// TIA Portal project "Respirator2020_V16" (V16) (continued)
REGION Network 5: Peep Supervisor
   RUNG wire#powerrail
      "VariableSupervisor_DB_Peep"(SetpointIncrement := "OperatingParameters".PeepPBPlus, SetpointDecrement := "OperatingParameters".PeepPBMinus, Max := 50.0, Min := 3.0, SetpointMax := "OperatingParameters".PeepMax, SetpointMin := "OperatingParameters".PeepMin, InOutSetpoint := "OperatingParameters".PeepSetpoint, InOutAlarmHI := "ProcessData".PeepSetpointAlarmHI, InOutPreAlarmHI := "ProcessData".PeepSetpointPreAlarmHI, InOutAlarmLOW := "ProcessData".PeepSetpointAlarmLOW, InOutPreAlarmLOW := "ProcessData".PeepSetpointPreAlarmLOW)
   END_RUNG
   // the same network as SCL:
   "VariableSupervisor_DB_Peep"(SetpointIncrement := "OperatingParameters".PeepPBPlus,   // "VariableSupervisor"
                           SetpointDecrement := "OperatingParameters".PeepPBMinus,
                           Max := 50.0,
                           Min := 3.0,
                           SetpointMax := "OperatingParameters".PeepMax,
                           SetpointMin := "OperatingParameters".PeepMin,
                           InOutSetpoint := "OperatingParameters".PeepSetpoint,
                           InOutAlarmHI := "ProcessData".PeepSetpointAlarmHI,
                           InOutPreAlarmHI := "ProcessData".PeepSetpointPreAlarmHI,
                           InOutAlarmLOW := "ProcessData".PeepSetpointAlarmLOW,
                           InOutPreAlarmLOW := "ProcessData".PeepSetpointPreAlarmLOW);
END_REGION

REGION Network 6: Frequency Supervisor
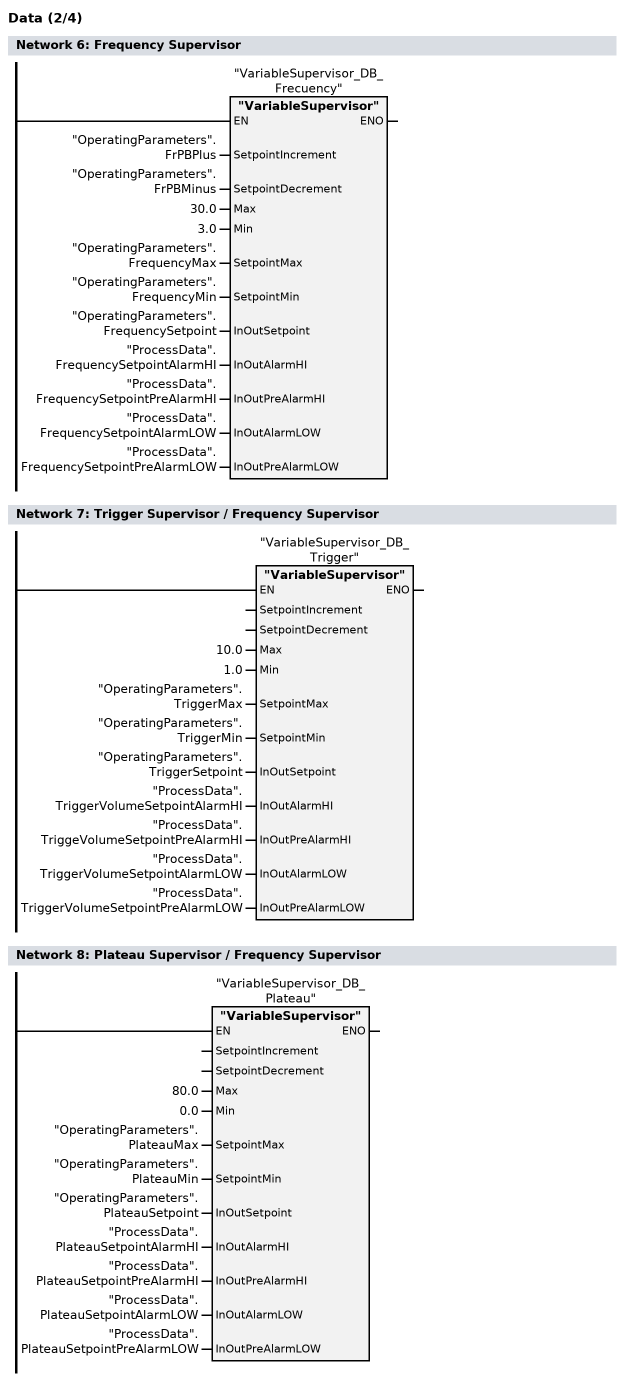
   RUNG wire#powerrail
      "VariableSupervisor_DB_Frecuency"(SetpointIncrement := "OperatingParameters".FrPBPlus, SetpointDecrement := "OperatingParameters".FrPBMinus, Max := 30.0, Min := 3.0, SetpointMax := "OperatingParameters".FrequencyMax, SetpointMin := "OperatingParameters".FrequencyMin, InOutSetpoint := "OperatingParameters".FrequencySetpoint, InOutAlarmHI := "ProcessData".FrequencySetpointAlarmHI, InOutPreAlarmHI := "ProcessData".FrequencySetpointPreAlarmHI, InOutAlarmLOW := "ProcessData".FrequencySetpointAlarmLOW, InOutPreAlarmLOW := "ProcessData".FrequencySetpointPreAlarmLOW)
   END_RUNG
   // the same network as SCL:
   "VariableSupervisor_DB_Frecuency"(SetpointIncrement := "OperatingParameters".FrPBPlus,   // "VariableSupervisor"
                           SetpointDecrement := "OperatingParameters".FrPBMinus,
                           Max := 30.0,
                           Min := 3.0,
                           SetpointMax := "OperatingParameters".FrequencyMax,
                           SetpointMin := "OperatingParameters".FrequencyMin,
                           InOutSetpoint := "OperatingParameters".FrequencySetpoint,
                           InOutAlarmHI := "ProcessData".FrequencySetpointAlarmHI,
                           InOutPreAlarmHI := "ProcessData".FrequencySetpointPreAlarmHI,
                           InOutAlarmLOW := "ProcessData".FrequencySetpointAlarmLOW,
                           InOutPreAlarmLOW := "ProcessData".FrequencySetpointPreAlarmLOW);
END_REGION

REGION Network 7: Trigger Supervisor / Frequency Supervisor
   RUNG wire#powerrail
      "VariableSupervisor_DB_Trigger"(SetpointIncrement :=, SetpointDecrement :=, Max := 10.0, Min := 1.0, SetpointMax := "OperatingParameters".TriggerMax, SetpointMin := "OperatingParameters".TriggerMin, InOutSetpoint := "OperatingParameters".TriggerSetpoint, InOutAlarmHI := "ProcessData".TriggerVolumeSetpointAlarmHI, InOutPreAlarmHI := "ProcessData".TriggeVolumeSetpointPreAlarmHI, InOutAlarmLOW := "ProcessData".TriggerVolumeSetpointAlarmLOW, InOutPreAlarmLOW := "ProcessData".TriggerVolumeSetpointPreAlarmLOW)
   END_RUNG
   // the same network as SCL:
   "VariableSupervisor_DB_Trigger"(Max := 10.0,   // "VariableSupervisor"
                           Min := 1.0,
                           SetpointMax := "OperatingParameters".TriggerMax,
                           SetpointMin := "OperatingParameters".TriggerMin,
                           InOutSetpoint := "OperatingParameters".TriggerSetpoint,
                           InOutAlarmHI := "ProcessData".TriggerVolumeSetpointAlarmHI,
                           InOutPreAlarmHI := "ProcessData".TriggeVolumeSetpointPreAlarmHI,
                           InOutAlarmLOW := "ProcessData".TriggerVolumeSetpointAlarmLOW,
                           InOutPreAlarmLOW := "ProcessData".TriggerVolumeSetpointPreAlarmLOW);
END_REGION

REGION Network 8: Plateau Supervisor / Frequency Supervisor
   RUNG wire#powerrail
      "VariableSupervisor_DB_Plateau"(SetpointIncrement :=, SetpointDecrement :=, Max := 80.0, Min := 0.0, SetpointMax := "OperatingParameters".PlateauMax, SetpointMin := "OperatingParameters".PlateauMin, InOutSetpoint := "OperatingParameters".PlateauSetpoint, InOutAlarmHI := "ProcessData".PlateauSetpointAlarmHI, InOutPreAlarmHI := "ProcessData".PlateauSetpointPreAlarmHI, InOutAlarmLOW := "ProcessData".PlateauSetpointAlarmLOW, InOutPreAlarmLOW := "ProcessData".PlateauSetpointPreAlarmLOW)
   END_RUNG
   // the same network as SCL:
   "VariableSupervisor_DB_Plateau"(Max := 80.0,   // "VariableSupervisor"
                           Min := 0.0,
                           SetpointMax := "OperatingParameters".PlateauMax,
                           SetpointMin := "OperatingParameters".PlateauMin,
                           InOutSetpoint := "OperatingParameters".PlateauSetpoint,
                           InOutAlarmHI := "ProcessData".PlateauSetpointAlarmHI,
                           InOutPreAlarmHI := "ProcessData".PlateauSetpointPreAlarmHI,
                           InOutAlarmLOW := "ProcessData".PlateauSetpointAlarmLOW,
                           InOutPreAlarmLOW := "ProcessData".PlateauSetpointPreAlarmLOW);
END_REGION

REGION Network 9: TidalVolume Supervisor / Frequency Supervisor
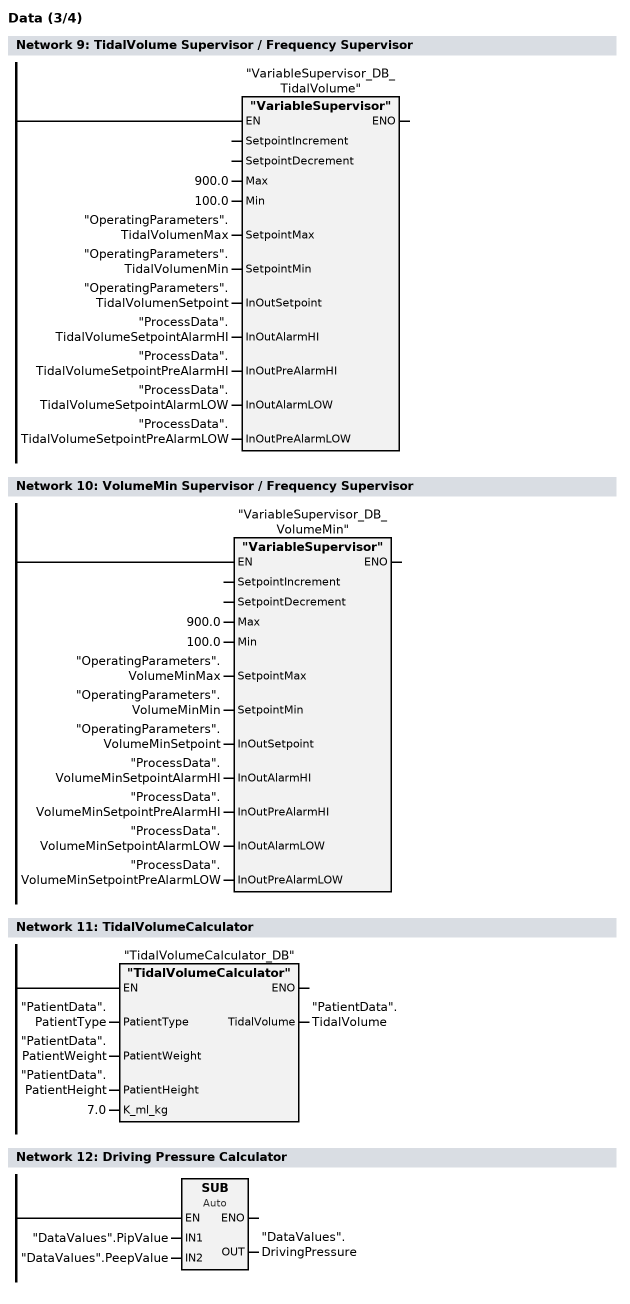
   RUNG wire#powerrail
      "VariableSupervisor_DB_TidalVolume"(SetpointIncrement :=, SetpointDecrement :=, Max := 900.0, Min := 100.0, SetpointMax := "OperatingParameters".TidalVolumenMax, SetpointMin := "OperatingParameters".TidalVolumenMin, InOutSetpoint := "OperatingParameters".TidalVolumenSetpoint, InOutAlarmHI := "ProcessData".TidalVolumeSetpointAlarmHI, InOutPreAlarmHI := "ProcessData".TidalVolumeSetpointPreAlarmHI, InOutAlarmLOW := "ProcessData".TidalVolumeSetpointAlarmLOW, InOutPreAlarmLOW := "ProcessData".TidalVolumeSetpointPreAlarmLOW)
   END_RUNG
   // the same network as SCL:
   "VariableSupervisor_DB_TidalVolume"(Max := 900.0,   // "VariableSupervisor"
                           Min := 100.0,
                           SetpointMax := "OperatingParameters".TidalVolumenMax,
                           SetpointMin := "OperatingParameters".TidalVolumenMin,
                           InOutSetpoint := "OperatingParameters".TidalVolumenSetpoint,
                           InOutAlarmHI := "ProcessData".TidalVolumeSetpointAlarmHI,
                           InOutPreAlarmHI := "ProcessData".TidalVolumeSetpointPreAlarmHI,
                           InOutAlarmLOW := "ProcessData".TidalVolumeSetpointAlarmLOW,
                           InOutPreAlarmLOW := "ProcessData".TidalVolumeSetpointPreAlarmLOW);
END_REGION

REGION Network 10: VolumeMin Supervisor / Frequency Supervisor
   RUNG wire#powerrail
      "VariableSupervisor_DB_VolumeMin"(SetpointIncrement :=, SetpointDecrement :=, Max := 900.0, Min := 100.0, SetpointMax := "OperatingParameters".VolumeMinMax, SetpointMin := "OperatingParameters".VolumeMinMin, InOutSetpoint := "OperatingParameters".VolumeMinSetpoint, InOutAlarmHI := "ProcessData".VolumeMinSetpointAlarmHI, InOutPreAlarmHI := "ProcessData".VolumeMinSetpointPreAlarmHI, InOutAlarmLOW := "ProcessData".VolumeMinSetpointAlarmLOW, InOutPreAlarmLOW := "ProcessData".VolumeMinSetpointPreAlarmLOW)
   END_RUNG
   // the same network as SCL:
   "VariableSupervisor_DB_VolumeMin"(Max := 900.0,   // "VariableSupervisor"
                           Min := 100.0,
                           SetpointMax := "OperatingParameters".VolumeMinMax,
                           SetpointMin := "OperatingParameters".VolumeMinMin,
                           InOutSetpoint := "OperatingParameters".VolumeMinSetpoint,
                           InOutAlarmHI := "ProcessData".VolumeMinSetpointAlarmHI,
                           InOutPreAlarmHI := "ProcessData".VolumeMinSetpointPreAlarmHI,
                           InOutAlarmLOW := "ProcessData".VolumeMinSetpointAlarmLOW,
                           InOutPreAlarmLOW := "ProcessData".VolumeMinSetpointPreAlarmLOW);
END_REGION

REGION Network 11: TidalVolumeCalculator
   RUNG wire#powerrail
      "TidalVolumeCalculator_DB"(PatientType := "PatientData".PatientType, PatientWeight := "PatientData".PatientWeight, PatientHeight := "PatientData".PatientHeight, K_ml_kg := 7.0, TidalVolume => "PatientData".TidalVolume)
   END_RUNG
   // the same network as SCL:
   "TidalVolumeCalculator_DB"(PatientType := "PatientData".PatientType,   // "TidalVolumeCalculator"
                           PatientWeight := "PatientData".PatientWeight,
                           PatientHeight := "PatientData".PatientHeight,
                           K_ml_kg := 7.0,
                           TidalVolume => "PatientData".TidalVolume);
END_REGION

REGION Network 12: Driving Pressure Calculator
   RUNG wire#powerrail
      Sub(in1 := "DataValues".PipValue, in2 := "DataValues".PeepValue, out => "DataValues".DrivingPressure)
   END_RUNG
   // the same network as SCL:
   "DataValues".DrivingPressure := "DataValues".PipValue - "DataValues".PeepValue;
END_REGION

REGION Network 13: Ratio Calculator
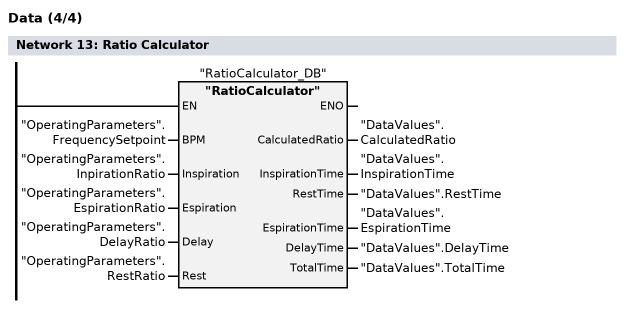
   RUNG wire#powerrail
      "RatioCalculator_DB"(BPM := "OperatingParameters".FrequencySetpoint, Inspiration := "OperatingParameters".InpirationRatio, Espiration := "OperatingParameters".EspirationRatio, Delay := "OperatingParameters".DelayRatio, Rest := "OperatingParameters".RestRatio, CalculatedRatio => "DataValues".CalculatedRatio, InspirationTime => "DataValues".InspirationTime, RestTime => "DataValues".RestTime, EspirationTime => "DataValues".EspirationTime, DelayTime => "DataValues".DelayTime, TotalTime => "DataValues".TotalTime)
   END_RUNG
   // the same network as SCL:
   "RatioCalculator_DB"(BPM := "OperatingParameters".FrequencySetpoint,   // "RatioCalculator"
                        Inspiration := "OperatingParameters".InpirationRatio,
                        Espiration := "OperatingParameters".EspirationRatio,
                        Delay := "OperatingParameters".DelayRatio,
                        Rest := "OperatingParameters".RestRatio,
                        CalculatedRatio => "DataValues".CalculatedRatio,
                        InspirationTime => "DataValues".InspirationTime,
                        RestTime => "DataValues".RestTime,
                        EspirationTime => "DataValues".EspirationTime,
                        DelayTime => "DataValues".DelayTime,
                        TotalTime => "DataValues".TotalTime);
END_REGION
END_FUNCTION_BLOCK

FUNCTION_BLOCK "TidalVolumeCalculator"   // FB11, SCL
{ S7_Optimized_Access := 'TRUE' }
AUTHOR : JL_Cristobal_2020
VERSION : 0.1
   VAR_INPUT
      PatientType : Int;
      PatientWeight : Real;
      PatientHeight : Real;
      K_ml_kg : Real;
   END_VAR
   VAR_OUTPUT
      TidalVolume : Real;
   END_VAR
   VAR
      CorrectedWeight : Real;
   END_VAR
BEGIN
   //**************************************************************************************************
   // TidalVolumeCalculator
   //**************************************************************************************************

   // Sex Selection
   CASE #PatientType OF
       1:  // Man
           #CorrectedWeight := 50.0;
       2:  // Woman
           #CorrectedWeight := 45.5;
       ELSE  // Not selected
           #CorrectedWeight := 0.0;;
   END_CASE;

   // Calc
   IF #CorrectedWeight <> 0 THEN
       #TidalVolume:= #K_ml_kg *((#CorrectedWeight+0.91)*(#PatientHeight));
       ELSE
           #TidalVolume := 0.0;
   END_IF;
END_FUNCTION_BLOCK

// folder: 2_SensorComm

FUNCTION_BLOCK "SensorComm_PtP_Freeport"   // FB20, SCL
{ S7_Optimized_Access := 'FALSE' }
AUTHOR : JL_Cristobal_2020
VERSION : 0.1
   VAR_OUTPUT
      OutputStatus : Struct
         Pressure1 : Real;
         Pressure2 : Real;
         VolumeAccumulated : Real;
         Flow : Real;
         TEMPERATURA_SONICA_PROMEDIO : Real;
         TEMPERATURA_PT100 : Real;
         HUMEDAD_RELATIVA : Real;
         PRESION_ATMOSFERICA : Real;
         DIRECCION_BRUJULA : Real;
         RADIACION_SOLAR : Real;
         VEL_PROMEDIO_VIENTO : Real;
         DIR_MEDIA_VIENTO : Real;
         HUMEDAD_ABSOLUTA : Real;
         PUNTO_ROCIO : Real;
         DIRECCION_VIENTO_GRADOS : Real;
         VEL_VIENTO_EJE_V : Real;
         VEL_VIENTO_EJE_U : Real;
         ERROR_MEDICION_VELOCIDAD : Bool;
         ERROR_MEDICION_BRUJULA : Bool;
         ERROR_MEDICION_TEMPERATURA : Bool;
         ERROR_MEDICION_HUMEDAD : Bool;
         ERROR_MEDICION_PRESION : Bool;
         ERROR_MEDICION_RADIACION_SOLAR : Bool;
      END_STRUCT;
      Pressure1 : Real;
      Pressure2 : Real;
      VolumeAccumulated : Real;
      Flow : Real;
      ErrorPressure1 : Bool;
      ErrorPressure2 : Bool;
      ErrorVolumeAccumulated : Bool;
      ErrorFlow : Bool;
   END_VAR
   VAR
      InputData : Struct
         Config_REQ : Bool;
         Reset_REQ : Bool;
      END_STRUCT;
      OutputData : Struct
         Config_DONE : Bool;
         Config_ERROR : Bool;
         Config_STAT : Word;
         Reset_DONE : Bool;
         Reset_ERROR : Bool;
         Reset_STAT : Word;
         Receive_P2P_NDR : Bool;
         Receive_P2P_ERROR : Bool;
         Receive_P2P_STAT : Word;
         Receive_P2P_Length : Word;
         Send_P2P_DONE : Bool;
         Send_P2P_ERROR : Bool;
         Send_P2P_STAT : Word;
      END_STRUCT;
      Control : Struct
         While_Section : Bool;
         COM_RST : Bool;
         Config_ERROR_save : Word;
         Reset_ERROR_save : Word;
         P2P_ERROR_save : Word;
         P2P_NDR_save : Word;
         Rcv_Length_save : Int;
      END_STRUCT;
      RecvBuffer : Array[1..254] of Byte;
      TransBuffer : Array[1..254] of Byte;
      IntermediateData : Struct
         Pressure1 : String;
         Pressure2 : String;
         VolumeAccumulated : String;
         Flow : String;
         Errors : String;
      END_STRUCT;
   END_VAR
BEGIN
   //**************************************************************************************************
   // Reading STATUS
   //**************************************************************************************************
   IF TRUE THEN
       // Pressure-1
       Chars_TO_Strg(Chars := "SensorComm_C_buffer_ptp".Ringbuffer,
                     pChars := 2,
                     Cnt := 6,
                     Strg => #IntermediateData.Pressure1);
       STRG_VAL(IN := #IntermediateData.Pressure1,
                FORMAT := W#16#0000,
                P := 1,
                OUT => #OutputStatus.Pressure1);
       #Pressure1 := #OutputStatus.Pressure1;

       // Pressure-2
       Chars_TO_Strg(Chars := "SensorComm_C_buffer_ptp".Ringbuffer,
                     pChars := 10,
                     Cnt := 6,
                     Strg => #IntermediateData.Pressure2);
       STRG_VAL(IN := #IntermediateData.Pressure2,
                FORMAT := W#16#0000,
                P := 1,
                OUT => #OutputStatus.Pressure2);
       #Pressure2 := #OutputStatus.Pressure2;

       // Volume Accumulated
       Chars_TO_Strg(Chars := "SensorComm_C_buffer_ptp".Ringbuffer,
                     pChars := 18,
                     Cnt := 6,
                     Strg => #IntermediateData.VolumeAccumulated);
       STRG_VAL(IN := #IntermediateData.VolumeAccumulated,
                FORMAT := W#16#0000,
                P := 1,
                OUT => #OutputStatus.VolumeAccumulated);
       #VolumeAccumulated := #OutputStatus.VolumeAccumulated;

       // Flow
       Chars_TO_Strg(Chars := "SensorComm_C_buffer_ptp".Ringbuffer,
                     pChars := 26,
                     Cnt := 6,
                     Strg => #IntermediateData.Flow);
       STRG_VAL(IN := #IntermediateData.Flow,
                FORMAT := W#16#0000,
                P := 1,
                OUT => #OutputStatus.Flow);
       #Flow := #OutputStatus.Flow;

        // Errors
       Chars_TO_Strg(Chars := "SensorComm_C_buffer_ptp".Ringbuffer,
                     pChars := 74,
                     Cnt := 6,
                     Strg => #IntermediateData.Errors);
   END_IF;
END_FUNCTION_BLOCK

// folder: 3_Alarms

FUNCTION_BLOCK "Alarms"   // FB5, LAD
TITLE = Alarms, Packing and Transport to HMI
{ S7_Optimized_Access := 'TRUE' }
AUTHOR : JL_Cristobal_2020
VERSION : 0.1
   VAR_IN_OUT
      AlarmsPack0 : Bool;
      AlarmsPack1 : Bool;
      AlarmsPack2 : Bool;
      AlarmsPack3 : Bool;
   END_VAR
BEGIN

REGION Network 1: Peak Alarms
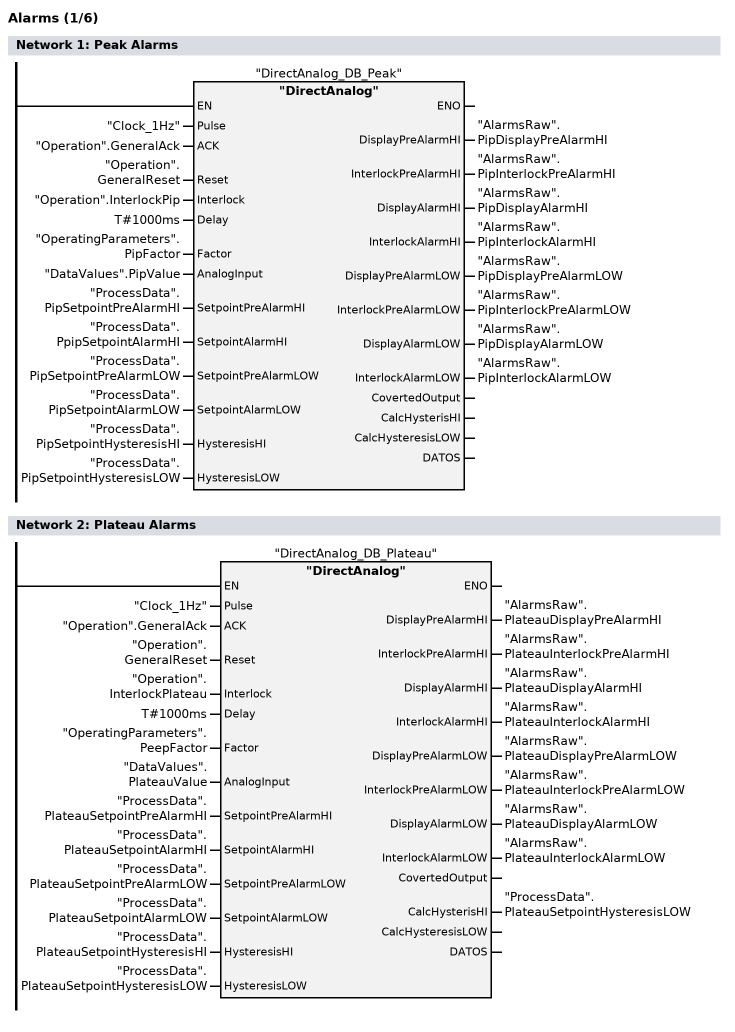
   RUNG wire#powerrail
      "DirectAnalog_DB_Peak"(Pulse := "Clock_1Hz", ACK := "Operation".GeneralAck, Reset := "Operation".GeneralReset, Interlock := "Operation".InterlockPip, Delay := T#1000ms, Factor := "OperatingParameters".PipFactor, AnalogInput := "DataValues".PipValue, SetpointPreAlarmHI := "ProcessData".PipSetpointPreAlarmHI, SetpointAlarmHI := "ProcessData".PpipSetpointAlarmHI, SetpointPreAlarmLOW := "ProcessData".PipSetpointPreAlarmLOW, SetpointAlarmLOW := "ProcessData".PipSetpointAlarmLOW, HysteresisHI := "ProcessData".PipSetpointHysteresisHI, HysteresisLOW := "ProcessData".PipSetpointHysteresisLOW, DisplayPreAlarmHI => "AlarmsRaw".PipDisplayPreAlarmHI, InterlockPreAlarmHI => "AlarmsRaw".PipInterlockPreAlarmHI, DisplayAlarmHI => "AlarmsRaw".PipDisplayAlarmHI, InterlockAlarmHI => "AlarmsRaw".PipInterlockAlarmHI, DisplayPreAlarmLOW => "AlarmsRaw".PipDisplayPreAlarmLOW, InterlockPreAlarmLOW => "AlarmsRaw".PipInterlockPreAlarmLOW, DisplayAlarmLOW => "AlarmsRaw".PipDisplayAlarmLOW, InterlockAlarmLOW => "AlarmsRaw".PipInterlockAlarmLOW, CovertedOutput =>, CalcHysterisHI =>, CalcHysteresisLOW =>, DATOS =>)
   END_RUNG
   // the same network as SCL:
   "DirectAnalog_DB_Peak"(Pulse := "Clock_1Hz",   // "DirectAnalog"
                          ACK := "Operation".GeneralAck,
                          Reset := "Operation".GeneralReset,
                          Interlock := "Operation".InterlockPip,
                          Delay := T#1000ms,
                          Factor := "OperatingParameters".PipFactor,
                          AnalogInput := "DataValues".PipValue,
                          SetpointPreAlarmHI := "ProcessData".PipSetpointPreAlarmHI,
                          SetpointAlarmHI := "ProcessData".PpipSetpointAlarmHI,
                          SetpointPreAlarmLOW := "ProcessData".PipSetpointPreAlarmLOW,
                          SetpointAlarmLOW := "ProcessData".PipSetpointAlarmLOW,
                          HysteresisHI := "ProcessData".PipSetpointHysteresisHI,
                          HysteresisLOW := "ProcessData".PipSetpointHysteresisLOW,
                          DisplayPreAlarmHI => "AlarmsRaw".PipDisplayPreAlarmHI,
                          InterlockPreAlarmHI => "AlarmsRaw".PipInterlockPreAlarmHI,
                          DisplayAlarmHI => "AlarmsRaw".PipDisplayAlarmHI,
                          InterlockAlarmHI => "AlarmsRaw".PipInterlockAlarmHI,
                          DisplayPreAlarmLOW => "AlarmsRaw".PipDisplayPreAlarmLOW,
                          InterlockPreAlarmLOW => "AlarmsRaw".PipInterlockPreAlarmLOW,
                          DisplayAlarmLOW => "AlarmsRaw".PipDisplayAlarmLOW,
                          InterlockAlarmLOW => "AlarmsRaw".PipInterlockAlarmLOW);
END_REGION

REGION Network 2: Plateau Alarms
   RUNG wire#powerrail
      "DirectAnalog_DB_Plateau"(Pulse := "Clock_1Hz", ACK := "Operation".GeneralAck, Reset := "Operation".GeneralReset, Interlock := "Operation".InterlockPlateau, Delay := T#1000ms, Factor := "OperatingParameters".PeepFactor, AnalogInput := "DataValues".PlateauValue, SetpointPreAlarmHI := "ProcessData".PlateauSetpointPreAlarmHI, SetpointAlarmHI := "ProcessData".PlateauSetpointAlarmHI, SetpointPreAlarmLOW := "ProcessData".PlateauSetpointPreAlarmLOW, SetpointAlarmLOW := "ProcessData".PlateauSetpointAlarmLOW, HysteresisHI := "ProcessData".PlateauSetpointHysteresisHI, HysteresisLOW := "ProcessData".PlateauSetpointHysteresisLOW, DisplayPreAlarmHI => "AlarmsRaw".PlateauDisplayPreAlarmHI, InterlockPreAlarmHI => "AlarmsRaw".PlateauInterlockPreAlarmHI, DisplayAlarmHI => "AlarmsRaw".PlateauDisplayAlarmHI, InterlockAlarmHI => "AlarmsRaw".PlateauInterlockAlarmHI, DisplayPreAlarmLOW => "AlarmsRaw".PlateauDisplayPreAlarmLOW, InterlockPreAlarmLOW => "AlarmsRaw".PlateauInterlockPreAlarmLOW, DisplayAlarmLOW => "AlarmsRaw".PlateauDisplayAlarmLOW, InterlockAlarmLOW => "AlarmsRaw".PlateauInterlockAlarmLOW, CovertedOutput =>, CalcHysterisHI => "ProcessData".PlateauSetpointHysteresisLOW, CalcHysteresisLOW =>, DATOS =>)
   END_RUNG
   // the same network as SCL:
   "DirectAnalog_DB_Plateau"(Pulse := "Clock_1Hz",   // "DirectAnalog"
                           ACK := "Operation".GeneralAck,
                           Reset := "Operation".GeneralReset,
                           Interlock := "Operation".InterlockPlateau,
                           Delay := T#1000ms,
                           Factor := "OperatingParameters".PeepFactor,
                           AnalogInput := "DataValues".PlateauValue,
                           SetpointPreAlarmHI := "ProcessData".PlateauSetpointPreAlarmHI,
                           SetpointAlarmHI := "ProcessData".PlateauSetpointAlarmHI,
                           SetpointPreAlarmLOW := "ProcessData".PlateauSetpointPreAlarmLOW,
                           SetpointAlarmLOW := "ProcessData".PlateauSetpointAlarmLOW,
                           HysteresisHI := "ProcessData".PlateauSetpointHysteresisHI,
                           HysteresisLOW := "ProcessData".PlateauSetpointHysteresisLOW,
                           DisplayPreAlarmHI => "AlarmsRaw".PlateauDisplayPreAlarmHI,
                           InterlockPreAlarmHI => "AlarmsRaw".PlateauInterlockPreAlarmHI,
                           DisplayAlarmHI => "AlarmsRaw".PlateauDisplayAlarmHI,
                           InterlockAlarmHI => "AlarmsRaw".PlateauInterlockAlarmHI,
                           DisplayPreAlarmLOW => "AlarmsRaw".PlateauDisplayPreAlarmLOW,
                           InterlockPreAlarmLOW => "AlarmsRaw".PlateauInterlockPreAlarmLOW,
                           DisplayAlarmLOW => "AlarmsRaw".PlateauDisplayAlarmLOW,
                           InterlockAlarmLOW => "AlarmsRaw".PlateauInterlockAlarmLOW,
                           CalcHysterisHI => "ProcessData".PlateauSetpointHysteresisLOW);
END_REGION

REGION Network 3: Peep Alarms
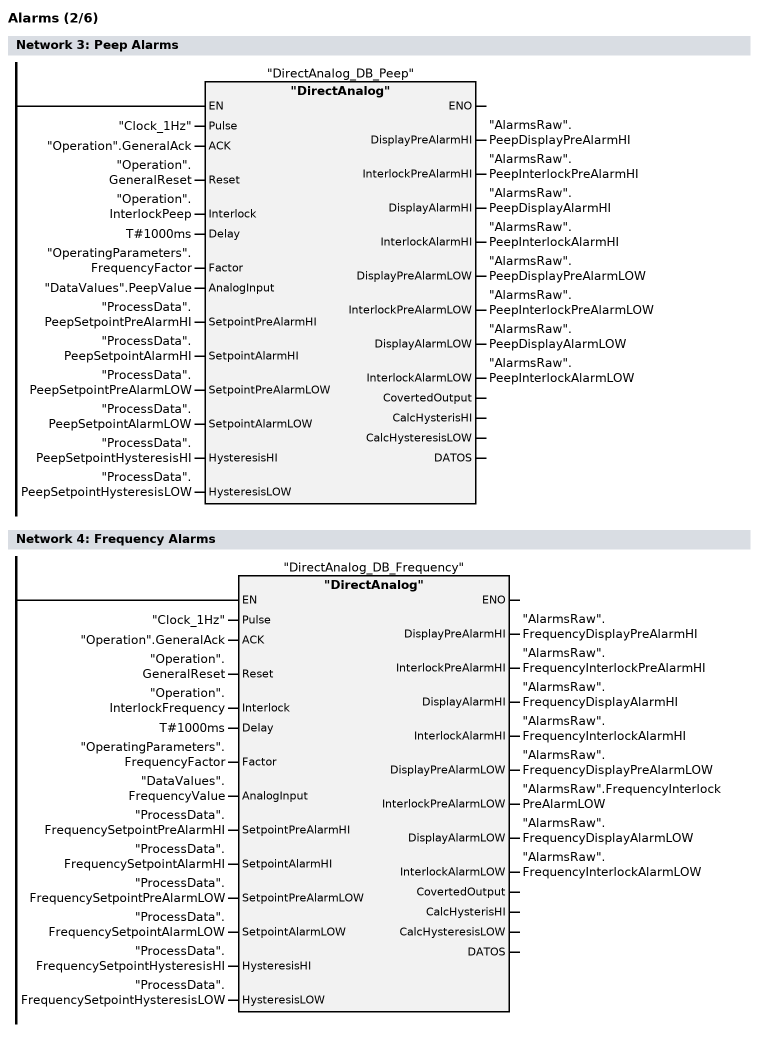
   RUNG wire#powerrail
      "DirectAnalog_DB_Peep"(Pulse := "Clock_1Hz", ACK := "Operation".GeneralAck, Reset := "Operation".GeneralReset, Interlock := "Operation".InterlockPeep, Delay := T#1000ms, Factor := "OperatingParameters".FrequencyFactor, AnalogInput := "DataValues".PeepValue, SetpointPreAlarmHI := "ProcessData".PeepSetpointPreAlarmHI, SetpointAlarmHI := "ProcessData".PeepSetpointAlarmHI, SetpointPreAlarmLOW := "ProcessData".PeepSetpointPreAlarmLOW, SetpointAlarmLOW := "ProcessData".PeepSetpointAlarmLOW, HysteresisHI := "ProcessData".PeepSetpointHysteresisHI, HysteresisLOW := "ProcessData".PeepSetpointHysteresisLOW, DisplayPreAlarmHI => "AlarmsRaw".PeepDisplayPreAlarmHI, InterlockPreAlarmHI => "AlarmsRaw".PeepInterlockPreAlarmHI, DisplayAlarmHI => "AlarmsRaw".PeepDisplayAlarmHI, InterlockAlarmHI => "AlarmsRaw".PeepInterlockAlarmHI, DisplayPreAlarmLOW => "AlarmsRaw".PeepDisplayPreAlarmLOW, InterlockPreAlarmLOW => "AlarmsRaw".PeepInterlockPreAlarmLOW, DisplayAlarmLOW => "AlarmsRaw".PeepDisplayAlarmLOW, InterlockAlarmLOW => "AlarmsRaw".PeepInterlockAlarmLOW, CovertedOutput =>, CalcHysterisHI =>, CalcHysteresisLOW =>, DATOS =>)
   END_RUNG
   // the same network as SCL:
   "DirectAnalog_DB_Peep"(Pulse := "Clock_1Hz",   // "DirectAnalog"
                          ACK := "Operation".GeneralAck,
                          Reset := "Operation".GeneralReset,
                          Interlock := "Operation".InterlockPeep,
                          Delay := T#1000ms,
                          Factor := "OperatingParameters".FrequencyFactor,
                          AnalogInput := "DataValues".PeepValue,
                          SetpointPreAlarmHI := "ProcessData".PeepSetpointPreAlarmHI,
                          SetpointAlarmHI := "ProcessData".PeepSetpointAlarmHI,
                          SetpointPreAlarmLOW := "ProcessData".PeepSetpointPreAlarmLOW,
                          SetpointAlarmLOW := "ProcessData".PeepSetpointAlarmLOW,
                          HysteresisHI := "ProcessData".PeepSetpointHysteresisHI,
                          HysteresisLOW := "ProcessData".PeepSetpointHysteresisLOW,
                          DisplayPreAlarmHI => "AlarmsRaw".PeepDisplayPreAlarmHI,
                          InterlockPreAlarmHI => "AlarmsRaw".PeepInterlockPreAlarmHI,
                          DisplayAlarmHI => "AlarmsRaw".PeepDisplayAlarmHI,
                          InterlockAlarmHI => "AlarmsRaw".PeepInterlockAlarmHI,
                          DisplayPreAlarmLOW => "AlarmsRaw".PeepDisplayPreAlarmLOW,
                          InterlockPreAlarmLOW => "AlarmsRaw".PeepInterlockPreAlarmLOW,
                          DisplayAlarmLOW => "AlarmsRaw".PeepDisplayAlarmLOW,
                          InterlockAlarmLOW => "AlarmsRaw".PeepInterlockAlarmLOW);
END_REGION

REGION Network 4: Frequency Alarms
   RUNG wire#powerrail
      "DirectAnalog_DB_Frequency"(Pulse := "Clock_1Hz", ACK := "Operation".GeneralAck, Reset := "Operation".GeneralReset, Interlock := "Operation".InterlockFrequency, Delay := T#1000ms, Factor := "OperatingParameters".FrequencyFactor, AnalogInput := "DataValues".FrequencyValue, SetpointPreAlarmHI := "ProcessData".FrequencySetpointPreAlarmHI, SetpointAlarmHI := "ProcessData".FrequencySetpointAlarmHI, SetpointPreAlarmLOW := "ProcessData".FrequencySetpointPreAlarmLOW, SetpointAlarmLOW := "ProcessData".FrequencySetpointAlarmLOW, HysteresisHI := "ProcessData".FrequencySetpointHysteresisHI, HysteresisLOW := "ProcessData".FrequencySetpointHysteresisLOW, DisplayPreAlarmHI => "AlarmsRaw".FrequencyDisplayPreAlarmHI, InterlockPreAlarmHI => "AlarmsRaw".FrequencyInterlockPreAlarmHI, DisplayAlarmHI => "AlarmsRaw".FrequencyDisplayAlarmHI, InterlockAlarmHI => "AlarmsRaw".FrequencyInterlockAlarmHI, DisplayPreAlarmLOW => "AlarmsRaw".FrequencyDisplayPreAlarmLOW, InterlockPreAlarmLOW => "AlarmsRaw".FrequencyInterlockPreAlarmLOW, DisplayAlarmLOW => "AlarmsRaw".FrequencyDisplayAlarmLOW, InterlockAlarmLOW => "AlarmsRaw".FrequencyInterlockAlarmLOW, CovertedOutput =>, CalcHysterisHI =>, CalcHysteresisLOW =>, DATOS =>)
   END_RUNG
   // the same network as SCL:
   "DirectAnalog_DB_Frequency"(Pulse := "Clock_1Hz",   // "DirectAnalog"
                           ACK := "Operation".GeneralAck,
                           Reset := "Operation".GeneralReset,
                           Interlock := "Operation".InterlockFrequency,
                           Delay := T#1000ms,
                           Factor := "OperatingParameters".FrequencyFactor,
                           AnalogInput := "DataValues".FrequencyValue,
                           SetpointPreAlarmHI := "ProcessData".FrequencySetpointPreAlarmHI,
                           SetpointAlarmHI := "ProcessData".FrequencySetpointAlarmHI,
                           SetpointPreAlarmLOW := "ProcessData".FrequencySetpointPreAlarmLOW,
                           SetpointAlarmLOW := "ProcessData".FrequencySetpointAlarmLOW,
                           HysteresisHI := "ProcessData".FrequencySetpointHysteresisHI,
                           HysteresisLOW := "ProcessData".FrequencySetpointHysteresisLOW,
                           DisplayPreAlarmHI => "AlarmsRaw".FrequencyDisplayPreAlarmHI,
                           InterlockPreAlarmHI => "AlarmsRaw".FrequencyInterlockPreAlarmHI,
                           DisplayAlarmHI => "AlarmsRaw".FrequencyDisplayAlarmHI,
                           InterlockAlarmHI => "AlarmsRaw".FrequencyInterlockAlarmHI,
                           DisplayPreAlarmLOW => "AlarmsRaw".FrequencyDisplayPreAlarmLOW,
                           InterlockPreAlarmLOW => "AlarmsRaw".FrequencyInterlockPreAlarmLOW,
                           DisplayAlarmLOW => "AlarmsRaw".FrequencyDisplayAlarmLOW,
                           InterlockAlarmLOW => "AlarmsRaw".FrequencyInterlockAlarmLOW);
END_REGION

REGION Network 5: Tidal Volume Alarms
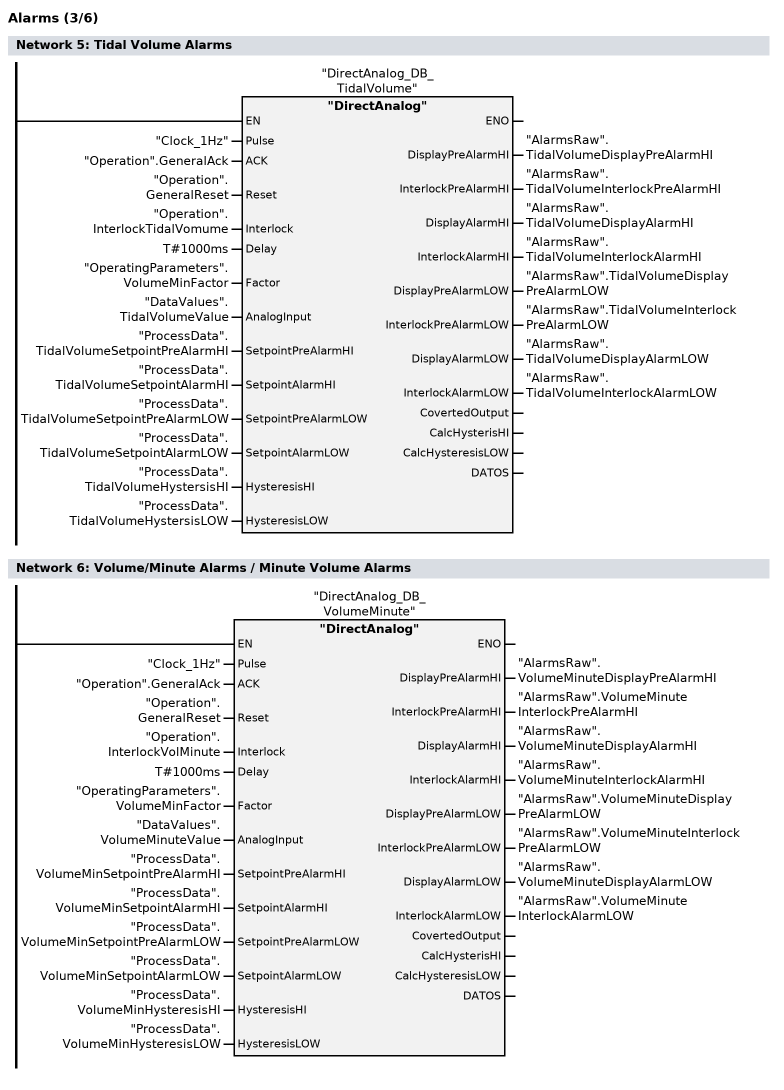
   RUNG wire#powerrail
      "DirectAnalog_DB_TidalVolume"(Pulse := "Clock_1Hz", ACK := "Operation".GeneralAck, Reset := "Operation".GeneralReset, Interlock := "Operation".InterlockTidalVomume, Delay := T#1000ms, Factor := "OperatingParameters".VolumeMinFactor, AnalogInput := "DataValues".TidalVolumeValue, SetpointPreAlarmHI := "ProcessData".TidalVolumeSetpointPreAlarmHI, SetpointAlarmHI := "ProcessData".TidalVolumeSetpointAlarmHI, SetpointPreAlarmLOW := "ProcessData".TidalVolumeSetpointPreAlarmLOW, SetpointAlarmLOW := "ProcessData".TidalVolumeSetpointAlarmLOW, HysteresisHI := "ProcessData".TidalVolumeHystersisHI, HysteresisLOW := "ProcessData".TidalVolumeHystersisLOW, DisplayPreAlarmHI => "AlarmsRaw".TidalVolumeDisplayPreAlarmHI, InterlockPreAlarmHI => "AlarmsRaw".TidalVolumeInterlockPreAlarmHI, DisplayAlarmHI => "AlarmsRaw".TidalVolumeDisplayAlarmHI, InterlockAlarmHI => "AlarmsRaw".TidalVolumeInterlockAlarmHI, DisplayPreAlarmLOW => "AlarmsRaw".TidalVolumeDisplayPreAlarmLOW, InterlockPreAlarmLOW => "AlarmsRaw".TidalVolumeInterlockPreAlarmLOW, DisplayAlarmLOW => "AlarmsRaw".TidalVolumeDisplayAlarmLOW, InterlockAlarmLOW => "AlarmsRaw".TidalVolumeInterlockAlarmLOW, CovertedOutput =>, CalcHysterisHI =>, CalcHysteresisLOW =>, DATOS =>)
   END_RUNG
   // the same network as SCL:
   "DirectAnalog_DB_TidalVolume"(Pulse := "Clock_1Hz",   // "DirectAnalog"
                           ACK := "Operation".GeneralAck,
                           Reset := "Operation".GeneralReset,
                           Interlock := "Operation".InterlockTidalVomume,
                           Delay := T#1000ms,
                           Factor := "OperatingParameters".VolumeMinFactor,
                           AnalogInput := "DataValues".TidalVolumeValue,
                           SetpointPreAlarmHI := "ProcessData".TidalVolumeSetpointPreAlarmHI,
                           SetpointAlarmHI := "ProcessData".TidalVolumeSetpointAlarmHI,
                           SetpointPreAlarmLOW := "ProcessData".TidalVolumeSetpointPreAlarmLOW,
                           SetpointAlarmLOW := "ProcessData".TidalVolumeSetpointAlarmLOW,
                           HysteresisHI := "ProcessData".TidalVolumeHystersisHI,
                           HysteresisLOW := "ProcessData".TidalVolumeHystersisLOW,
                           DisplayPreAlarmHI => "AlarmsRaw".TidalVolumeDisplayPreAlarmHI,
                           InterlockPreAlarmHI => "AlarmsRaw".TidalVolumeInterlockPreAlarmHI,
                           DisplayAlarmHI => "AlarmsRaw".TidalVolumeDisplayAlarmHI,
                           InterlockAlarmHI => "AlarmsRaw".TidalVolumeInterlockAlarmHI,
                           DisplayPreAlarmLOW => "AlarmsRaw".TidalVolumeDisplayPreAlarmLOW,
                           InterlockPreAlarmLOW => "AlarmsRaw".TidalVolumeInterlockPreAlarmLOW,
                           DisplayAlarmLOW => "AlarmsRaw".TidalVolumeDisplayAlarmLOW,
                           InterlockAlarmLOW => "AlarmsRaw".TidalVolumeInterlockAlarmLOW);
END_REGION
